REGION Network 5: Estado 3
   RUNG wire#powerrail
      { S7_Templates := "SrcType := DWord" } EQ_Contact(in1 := #Prioritaria, in2 := 16#0000_0000)
      { S7_Templates := "SrcType := DWord" } EQ_Contact(in1 := #Concatenadora, in2 := 16#0000_0004)
      wire#w1
      I_Contact( #"Falla Prioritarias" )
      I_Contact( #"Error Concatenadoras" )
      { S7_GenerateENO := "TRUE" } Move(in := 16#0000_0004, out1 => #Estado)
   END_RUNG
   RUNG wire#powerrail
      { S7_Templates := "SrcType := DWord" } EQ_Contact(in1 := #Prioritaria, in2 := 16#0000_0004)
   END_RUNG wire#w1
   // the same network as SCL:
   IF (((#Prioritaria = 16#0000_0000) AND (#Concatenadora = 16#0000_0004)) OR (#Prioritaria = 16#0000_0004)) AND NOT #"Falla Prioritarias" AND NOT #"Error Concatenadoras" THEN
       #Estado := 16#0000_0004;
   END_IF;
END_REGION

REGION Network 6: Estado 4
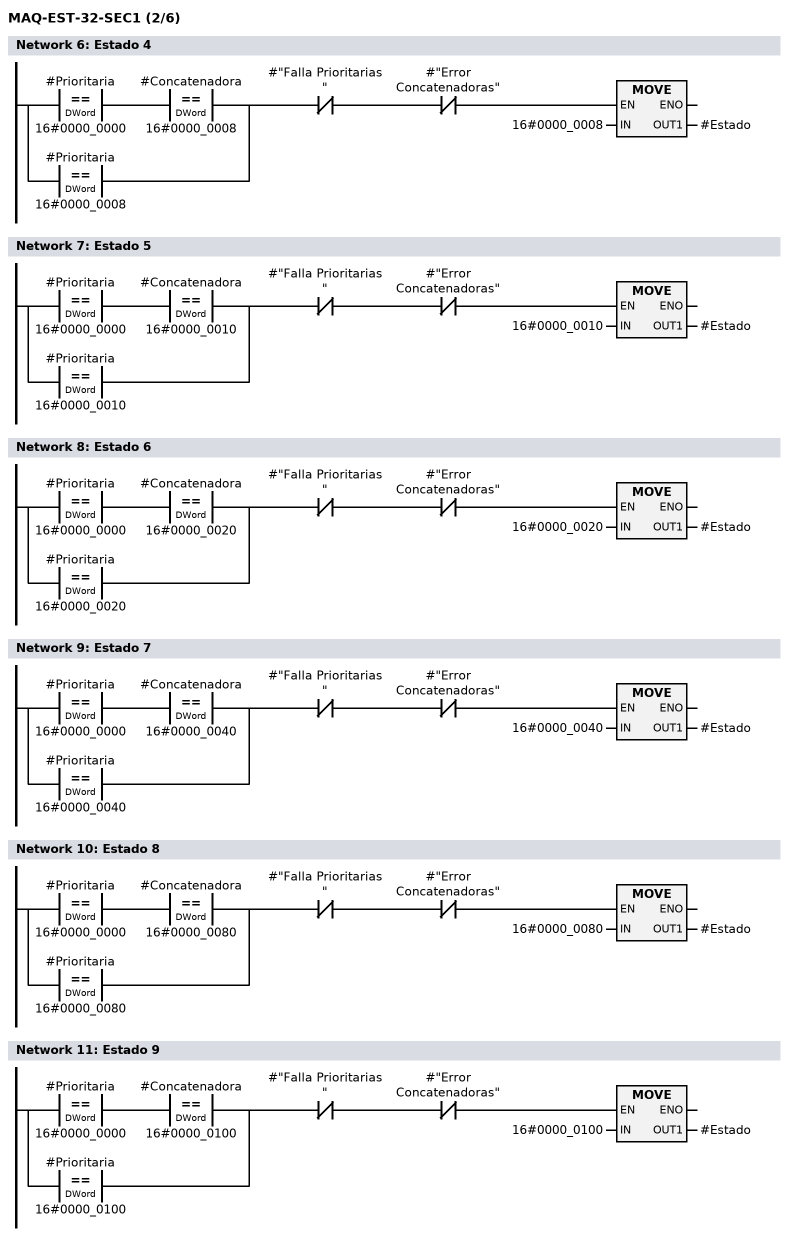
   RUNG wire#powerrail
      { S7_Templates := "SrcType := DWord" } EQ_Contact(in1 := #Prioritaria, in2 := 16#0000_0000)
      { S7_Templates := "SrcType := DWord" } EQ_Contact(in1 := #Concatenadora, in2 := 16#0000_0008)
      wire#w1
      I_Contact( #"Falla Prioritarias" )
      I_Contact( #"Error Concatenadoras" )
      { S7_GenerateENO := "TRUE" } Move(in := 16#0000_0008, out1 => #Estado)
   END_RUNG
   RUNG wire#powerrail
      { S7_Templates := "SrcType := DWord" } EQ_Contact(in1 := #Prioritaria, in2 := 16#0000_0008)
   END_RUNG wire#w1
   // the same network as SCL:
   IF (((#Prioritaria = 16#0000_0000) AND (#Concatenadora = 16#0000_0008)) OR (#Prioritaria = 16#0000_0008)) AND NOT #"Falla Prioritarias" AND NOT #"Error Concatenadoras" THEN
       #Estado := 16#0000_0008;
   END_IF;
END_REGION

REGION Network 7: Estado 5
   RUNG wire#powerrail
      { S7_Templates := "SrcType := DWord" } EQ_Contact(in1 := #Prioritaria, in2 := 16#0000_0000)
      { S7_Templates := "SrcType := DWord" } EQ_Contact(in1 := #Concatenadora, in2 := 16#0000_0010)
      wire#w1
      I_Contact( #"Falla Prioritarias" )
      I_Contact( #"Error Concatenadoras" )
      { S7_GenerateENO := "TRUE" } Move(in := 16#0000_0010, out1 => #Estado)
   END_RUNG
   RUNG wire#powerrail
      { S7_Templates := "SrcType := DWord" } EQ_Contact(in1 := #Prioritaria, in2 := 16#0000_0010)
   END_RUNG wire#w1
   // the same network as SCL:
   IF (((#Prioritaria = 16#0000_0000) AND (#Concatenadora = 16#0000_0010)) OR (#Prioritaria = 16#0000_0010)) AND NOT #"Falla Prioritarias" AND NOT #"Error Concatenadoras" THEN
       #Estado := 16#0000_0010;
   END_IF;
END_REGION

REGION Network 8: Estado 6
   RUNG wire#powerrail
      { S7_Templates := "SrcType := DWord" } EQ_Contact(in1 := #Prioritaria, in2 := 16#0000_0000)
      { S7_Templates := "SrcType := DWord" } EQ_Contact(in1 := #Concatenadora, in2 := 16#0000_0020)
      wire#w1
      I_Contact( #"Falla Prioritarias" )
      I_Contact( #"Error Concatenadoras" )
      { S7_GenerateENO := "TRUE" } Move(in := 16#0000_0020, out1 => #Estado)
   END_RUNG
   RUNG wire#powerrail
      { S7_Templates := "SrcType := DWord" } EQ_Contact(in1 := #Prioritaria, in2 := 16#0000_0020)
   END_RUNG wire#w1
   // the same network as SCL:
   IF (((#Prioritaria = 16#0000_0000) AND (#Concatenadora = 16#0000_0020)) OR (#Prioritaria = 16#0000_0020)) AND NOT #"Falla Prioritarias" AND NOT #"Error Concatenadoras" THEN
       #Estado := 16#0000_0020;
   END_IF;
END_REGION

REGION Network 9: Estado 7
   RUNG wire#powerrail
      { S7_Templates := "SrcType := DWord" } EQ_Contact(in1 := #Prioritaria, in2 := 16#0000_0000)
      { S7_Templates := "SrcType := DWord" } EQ_Contact(in1 := #Concatenadora, in2 := 16#0000_0040)
      wire#w1
      I_Contact( #"Falla Prioritarias" )
      I_Contact( #"Error Concatenadoras" )
      { S7_GenerateENO := "TRUE" } Move(in := 16#0000_0040, out1 => #Estado)
   END_RUNG
   RUNG wire#powerrail
      { S7_Templates := "SrcType := DWord" } EQ_Contact(in1 := #Prioritaria, in2 := 16#0000_0040)
   END_RUNG wire#w1
   // the same network as SCL:
   IF (((#Prioritaria = 16#0000_0000) AND (#Concatenadora = 16#0000_0040)) OR (#Prioritaria = 16#0000_0040)) AND NOT #"Falla Prioritarias" AND NOT #"Error Concatenadoras" THEN
       #Estado := 16#0000_0040;
   END_IF;
END_REGION

REGION Network 10: Estado 8
   RUNG wire#powerrail
      { S7_Templates := "SrcType := DWord" } EQ_Contact(in1 := #Prioritaria, in2 := 16#0000_0000)
      { S7_Templates := "SrcType := DWord" } EQ_Contact(in1 := #Concatenadora, in2 := 16#0000_0080)
      wire#w1
      I_Contact( #"Falla Prioritarias" )
      I_Contact( #"Error Concatenadoras" )
      { S7_GenerateENO := "TRUE" } Move(in := 16#0000_0080, out1 => #Estado)
   END_RUNG
   RUNG wire#powerrail
      { S7_Templates := "SrcType := DWord" } EQ_Contact(in1 := #Prioritaria, in2 := 16#0000_0080)
   END_RUNG wire#w1
   // the same network as SCL:
   IF (((#Prioritaria = 16#0000_0000) AND (#Concatenadora = 16#0000_0080)) OR (#Prioritaria = 16#0000_0080)) AND NOT #"Falla Prioritarias" AND NOT #"Error Concatenadoras" THEN
       #Estado := 16#0000_0080;
   END_IF;
END_REGION

REGION Network 11: Estado 9
   RUNG wire#powerrail
      { S7_Templates := "SrcType := DWord" } EQ_Contact(in1 := #Prioritaria, in2 := 16#0000_0000)
      { S7_Templates := "SrcType := DWord" } EQ_Contact(in1 := #Concatenadora, in2 := 16#0000_0100)
      wire#w1
      I_Contact( #"Falla Prioritarias" )
      I_Contact( #"Error Concatenadoras" )
      { S7_GenerateENO := "TRUE" } Move(in := 16#0000_0100, out1 => #Estado)
   END_RUNG
   RUNG wire#powerrail
      { S7_Templates := "SrcType := DWord" } EQ_Contact(in1 := #Prioritaria, in2 := 16#0000_0100)
   END_RUNG wire#w1
   // the same network as SCL:
   IF (((#Prioritaria = 16#0000_0000) AND (#Concatenadora = 16#0000_0100)) OR (#Prioritaria = 16#0000_0100)) AND NOT #"Falla Prioritarias" AND NOT #"Error Concatenadoras" THEN
       #Estado := 16#0000_0100;
   END_IF;
END_REGION

REGION Network 12: Estado 10
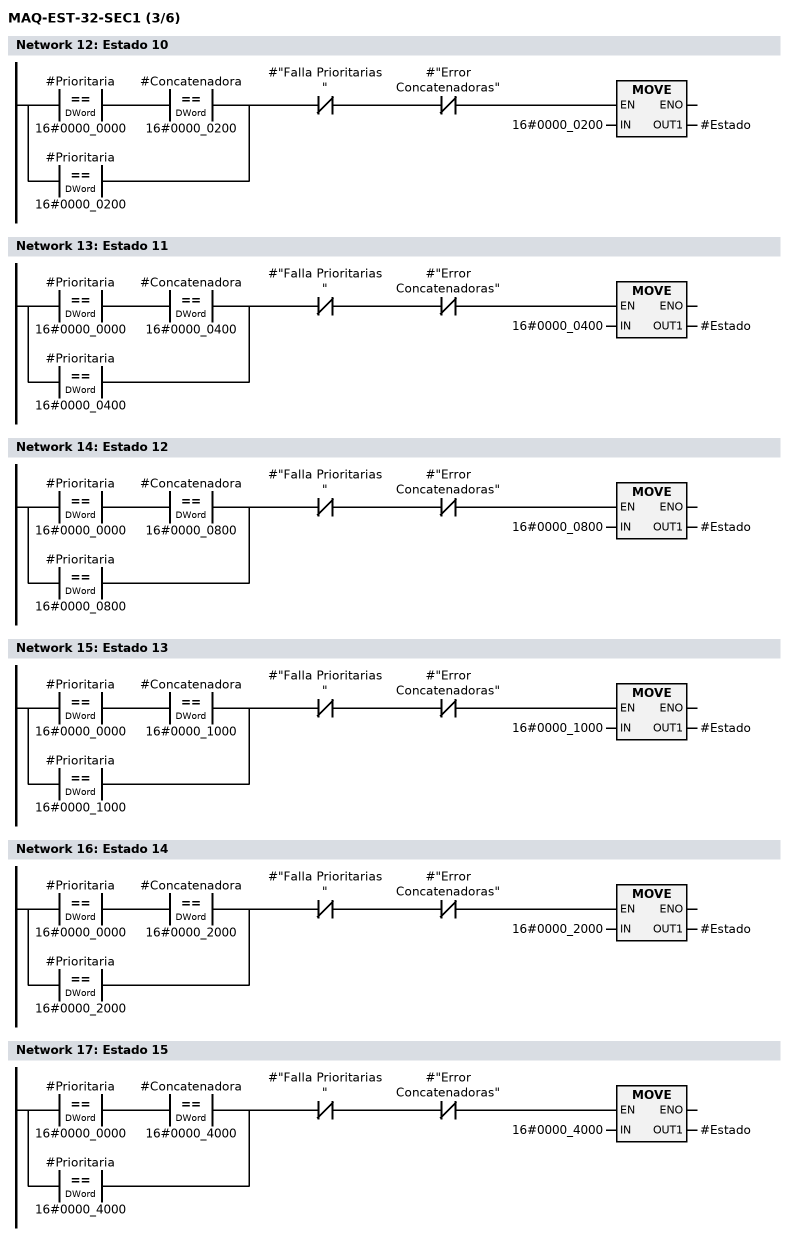
   RUNG wire#powerrail
      { S7_Templates := "SrcType := DWord" } EQ_Contact(in1 := #Prioritaria, in2 := 16#0000_0000)
      { S7_Templates := "SrcType := DWord" } EQ_Contact(in1 := #Concatenadora, in2 := 16#0000_0200)
      wire#w1
      I_Contact( #"Falla Prioritarias" )
      I_Contact( #"Error Concatenadoras" )
      { S7_GenerateENO := "TRUE" } Move(in := 16#0000_0200, out1 => #Estado)
   END_RUNG
   RUNG wire#powerrail
      { S7_Templates := "SrcType := DWord" } EQ_Contact(in1 := #Prioritaria, in2 := 16#0000_0200)
   END_RUNG wire#w1
   // the same network as SCL:
   IF (((#Prioritaria = 16#0000_0000) AND (#Concatenadora = 16#0000_0200)) OR (#Prioritaria = 16#0000_0200)) AND NOT #"Falla Prioritarias" AND NOT #"Error Concatenadoras" THEN
       #Estado := 16#0000_0200;
   END_IF;
END_REGION

REGION Network 13: Estado 11
   RUNG wire#powerrail
      { S7_Templates := "SrcType := DWord" } EQ_Contact(in1 := #Prioritaria, in2 := 16#0000_0000)
      { S7_Templates := "SrcType := DWord" } EQ_Contact(in1 := #Concatenadora, in2 := 16#0000_0400)
      wire#w1
      I_Contact( #"Falla Prioritarias" )
      I_Contact( #"Error Concatenadoras" )
      { S7_GenerateENO := "TRUE" } Move(in := 16#0000_0400, out1 => #Estado)
   END_RUNG
   RUNG wire#powerrail
      { S7_Templates := "SrcType := DWord" } EQ_Contact(in1 := #Prioritaria, in2 := 16#0000_0400)
   END_RUNG wire#w1
   // the same network as SCL:
   IF (((#Prioritaria = 16#0000_0000) AND (#Concatenadora = 16#0000_0400)) OR (#Prioritaria = 16#0000_0400)) AND NOT #"Falla Prioritarias" AND NOT #"Error Concatenadoras" THEN
       #Estado := 16#0000_0400;
   END_IF;
END_REGION

REGION Network 14: Estado 12
   RUNG wire#powerrail
      { S7_Templates := "SrcType := DWord" } EQ_Contact(in1 := #Prioritaria, in2 := 16#0000_0000)
      { S7_Templates := "SrcType := DWord" } EQ_Contact(in1 := #Concatenadora, in2 := 16#0000_0800)
      wire#w1
      I_Contact( #"Falla Prioritarias" )
      I_Contact( #"Error Concatenadoras" )
      { S7_GenerateENO := "TRUE" } Move(in := 16#0000_0800, out1 => #Estado)
   END_RUNG
   RUNG wire#powerrail
      { S7_Templates := "SrcType := DWord" } EQ_Contact(in1 := #Prioritaria, in2 := 16#0000_0800)
   END_RUNG wire#w1
   // the same network as SCL:
   IF (((#Prioritaria = 16#0000_0000) AND (#Concatenadora = 16#0000_0800)) OR (#Prioritaria = 16#0000_0800)) AND NOT #"Falla Prioritarias" AND NOT #"Error Concatenadoras" THEN
       #Estado := 16#0000_0800;
   END_IF;
END_REGION

REGION Network 15: Estado 13
   RUNG wire#powerrail
      { S7_Templates := "SrcType := DWord" } EQ_Contact(in1 := #Prioritaria, in2 := 16#0000_0000)
      { S7_Templates := "SrcType := DWord" } EQ_Contact(in1 := #Concatenadora, in2 := 16#0000_1000)
      wire#w1
      I_Contact( #"Falla Prioritarias" )
      I_Contact( #"Error Concatenadoras" )
      { S7_GenerateENO := "TRUE" } Move(in := 16#0000_1000, out1 => #Estado)
   END_RUNG
   RUNG wire#powerrail
      { S7_Templates := "SrcType := DWord" } EQ_Contact(in1 := #Prioritaria, in2 := 16#0000_1000)
   END_RUNG wire#w1
   // the same network as SCL:
   IF (((#Prioritaria = 16#0000_0000) AND (#Concatenadora = 16#0000_1000)) OR (#Prioritaria = 16#0000_1000)) AND NOT #"Falla Prioritarias" AND NOT #"Error Concatenadoras" THEN
       #Estado := 16#0000_1000;
   END_IF;
END_REGION

REGION Network 16: Estado 14
   RUNG wire#powerrail
      { S7_Templates := "SrcType := DWord" } EQ_Contact(in1 := #Prioritaria, in2 := 16#0000_0000)
      { S7_Templates := "SrcType := DWord" } EQ_Contact(in1 := #Concatenadora, in2 := 16#0000_2000)
      wire#w1
      I_Contact( #"Falla Prioritarias" )
      I_Contact( #"Error Concatenadoras" )
      { S7_GenerateENO := "TRUE" } Move(in := 16#0000_2000, out1 => #Estado)
   END_RUNG
   RUNG wire#powerrail
      { S7_Templates := "SrcType := DWord" } EQ_Contact(in1 := #Prioritaria, in2 := 16#0000_2000)
   END_RUNG wire#w1
   // the same network as SCL:
   IF (((#Prioritaria = 16#0000_0000) AND (#Concatenadora = 16#0000_2000)) OR (#Prioritaria = 16#0000_2000)) AND NOT #"Falla Prioritarias" AND NOT #"Error Concatenadoras" THEN
       #Estado := 16#0000_2000;
   END_IF;
END_REGION

REGION Network 17: Estado 15
   RUNG wire#powerrail
      { S7_Templates := "SrcType := DWord" } EQ_Contact(in1 := #Prioritaria, in2 := 16#0000_0000)
      { S7_Templates := "SrcType := DWord" } EQ_Contact(in1 := #Concatenadora, in2 := 16#0000_4000)
      wire#w1
      I_Contact( #"Falla Prioritarias" )
      I_Contact( #"Error Concatenadoras" )
      { S7_GenerateENO := "TRUE" } Move(in := 16#0000_4000, out1 => #Estado)
   END_RUNG
   RUNG wire#powerrail
      { S7_Templates := "SrcType := DWord" } EQ_Contact(in1 := #Prioritaria, in2 := 16#0000_4000)
   END_RUNG wire#w1
   // the same network as SCL:
   IF (((#Prioritaria = 16#0000_0000) AND (#Concatenadora = 16#0000_4000)) OR (#Prioritaria = 16#0000_4000)) AND NOT #"Falla Prioritarias" AND NOT #"Error Concatenadoras" THEN
       #Estado := 16#0000_4000;
   END_IF;
END_REGION

REGION Network 18: Estado 16
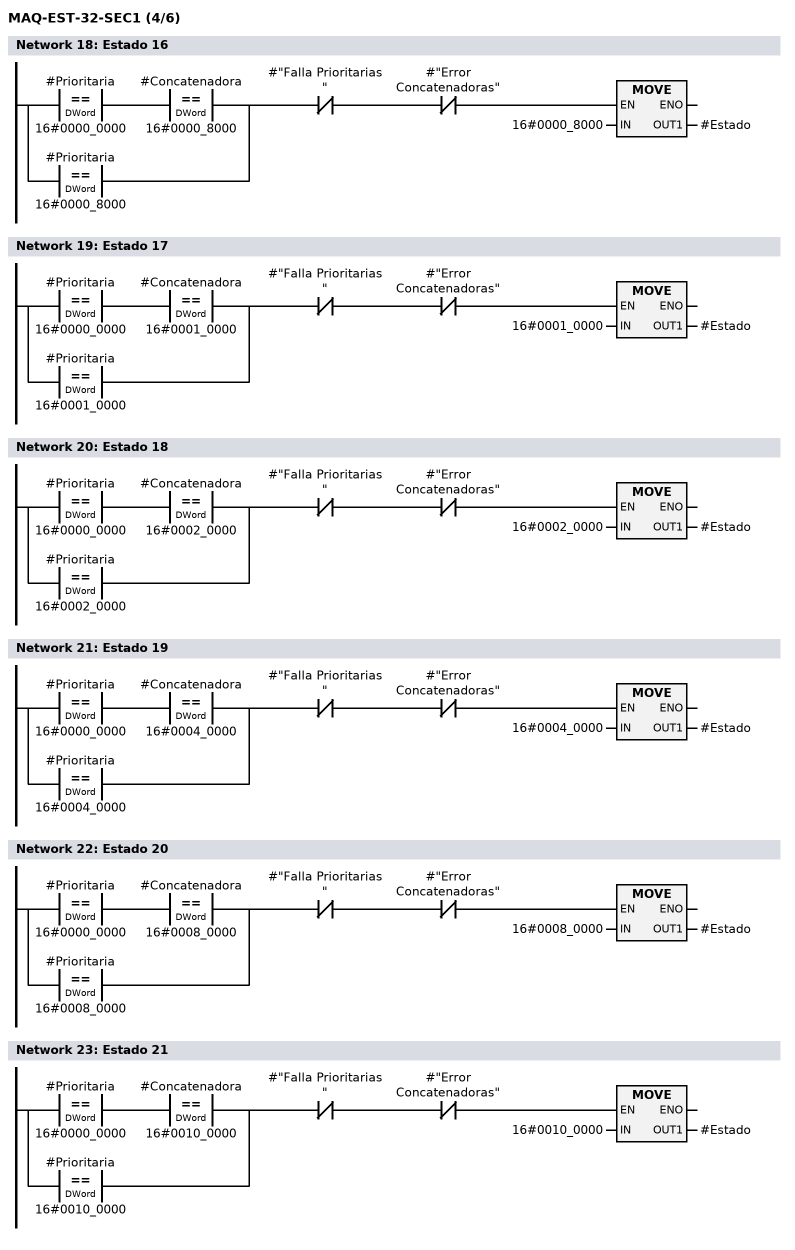
   RUNG wire#powerrail
      { S7_Templates := "SrcType := DWord" } EQ_Contact(in1 := #Prioritaria, in2 := 16#0000_0000)
      { S7_Templates := "SrcType := DWord" } EQ_Contact(in1 := #Concatenadora, in2 := 16#0000_8000)
      wire#w1
      I_Contact( #"Falla Prioritarias" )
      I_Contact( #"Error Concatenadoras" )
      { S7_GenerateENO := "TRUE" } Move(in := 16#0000_8000, out1 => #Estado)
   END_RUNG
   RUNG wire#powerrail
      { S7_Templates := "SrcType := DWord" } EQ_Contact(in1 := #Prioritaria, in2 := 16#0000_8000)
   END_RUNG wire#w1
   // the same network as SCL:
   IF (((#Prioritaria = 16#0000_0000) AND (#Concatenadora = 16#0000_8000)) OR (#Prioritaria = 16#0000_8000)) AND NOT #"Falla Prioritarias" AND NOT #"Error Concatenadoras" THEN
       #Estado := 16#0000_8000;
   END_IF;
END_REGION

REGION Network 19: Estado 17
   RUNG wire#powerrail
      { S7_Templates := "SrcType := DWord" } EQ_Contact(in1 := #Prioritaria, in2 := 16#0000_0000)
      { S7_Templates := "SrcType := DWord" } EQ_Contact(in1 := #Concatenadora, in2 := 16#0001_0000)
      wire#w1
      I_Contact( #"Falla Prioritarias" )
      I_Contact( #"Error Concatenadoras" )
      { S7_GenerateENO := "TRUE" } Move(in := 16#0001_0000, out1 => #Estado)
   END_RUNG
   RUNG wire#powerrail
      { S7_Templates := "SrcType := DWord" } EQ_Contact(in1 := #Prioritaria, in2 := 16#0001_0000)
   END_RUNG wire#w1
   // the same network as SCL:
   IF (((#Prioritaria = 16#0000_0000) AND (#Concatenadora = 16#0001_0000)) OR (#Prioritaria = 16#0001_0000)) AND NOT #"Falla Prioritarias" AND NOT #"Error Concatenadoras" THEN
       #Estado := 16#0001_0000;
   END_IF;
END_REGION

REGION Network 20: Estado 18
   RUNG wire#powerrail
      { S7_Templates := "SrcType := DWord" } EQ_Contact(in1 := #Prioritaria, in2 := 16#0000_0000)
      { S7_Templates := "SrcType := DWord" } EQ_Contact(in1 := #Concatenadora, in2 := 16#0002_0000)
      wire#w1
      I_Contact( #"Falla Prioritarias" )
      I_Contact( #"Error Concatenadoras" )
      { S7_GenerateENO := "TRUE" } Move(in := 16#0002_0000, out1 => #Estado)
   END_RUNG
   RUNG wire#powerrail
      { S7_Templates := "SrcType := DWord" } EQ_Contact(in1 := #Prioritaria, in2 := 16#0002_0000)
   END_RUNG wire#w1
   // the same network as SCL:
   IF (((#Prioritaria = 16#0000_0000) AND (#Concatenadora = 16#0002_0000)) OR (#Prioritaria = 16#0002_0000)) AND NOT #"Falla Prioritarias" AND NOT #"Error Concatenadoras" THEN
       #Estado := 16#0002_0000;
   END_IF;
END_REGION

REGION Network 21: Estado 19
   RUNG wire#powerrail
      { S7_Templates := "SrcType := DWord" } EQ_Contact(in1 := #Prioritaria, in2 := 16#0000_0000)
      { S7_Templates := "SrcType := DWord" } EQ_Contact(in1 := #Concatenadora, in2 := 16#0004_0000)
      wire#w1
      I_Contact( #"Falla Prioritarias" )
      I_Contact( #"Error Concatenadoras" )
      { S7_GenerateENO := "TRUE" } Move(in := 16#0004_0000, out1 => #Estado)
   END_RUNG
   RUNG wire#powerrail
      { S7_Templates := "SrcType := DWord" } EQ_Contact(in1 := #Prioritaria, in2 := 16#0004_0000)
   END_RUNG wire#w1
   // the same network as SCL:
   IF (((#Prioritaria = 16#0000_0000) AND (#Concatenadora = 16#0004_0000)) OR (#Prioritaria = 16#0004_0000)) AND NOT #"Falla Prioritarias" AND NOT #"Error Concatenadoras" THEN
       #Estado := 16#0004_0000;
   END_IF;
END_REGION

REGION Network 22: Estado 20
   RUNG wire#powerrail
      { S7_Templates := "SrcType := DWord" } EQ_Contact(in1 := #Prioritaria, in2 := 16#0000_0000)
      { S7_Templates := "SrcType := DWord" } EQ_Contact(in1 := #Concatenadora, in2 := 16#0008_0000)
      wire#w1
      I_Contact( #"Falla Prioritarias" )
      I_Contact( #"Error Concatenadoras" )
      { S7_GenerateENO := "TRUE" } Move(in := 16#0008_0000, out1 => #Estado)
   END_RUNG
   RUNG wire#powerrail
      { S7_Templates := "SrcType := DWord" } EQ_Contact(in1 := #Prioritaria, in2 := 16#0008_0000)
   END_RUNG wire#w1
   // the same network as SCL:
   IF (((#Prioritaria = 16#0000_0000) AND (#Concatenadora = 16#0008_0000)) OR (#Prioritaria = 16#0008_0000)) AND NOT #"Falla Prioritarias" AND NOT #"Error Concatenadoras" THEN
       #Estado := 16#0008_0000;
   END_IF;
END_REGION

REGION Network 23: Estado 21
   RUNG wire#powerrail
      { S7_Templates := "SrcType := DWord" } EQ_Contact(in1 := #Prioritaria, in2 := 16#0000_0000)
      { S7_Templates := "SrcType := DWord" } EQ_Contact(in1 := #Concatenadora, in2 := 16#0010_0000)
      wire#w1
      I_Contact( #"Falla Prioritarias" )
      I_Contact( #"Error Concatenadoras" )
      { S7_GenerateENO := "TRUE" } Move(in := 16#0010_0000, out1 => #Estado)
   END_RUNG
   RUNG wire#powerrail
      { S7_Templates := "SrcType := DWord" } EQ_Contact(in1 := #Prioritaria, in2 := 16#0010_0000)
   END_RUNG wire#w1
   // the same network as SCL:
   IF (((#Prioritaria = 16#0000_0000) AND (#Concatenadora = 16#0010_0000)) OR (#Prioritaria = 16#0010_0000)) AND NOT #"Falla Prioritarias" AND NOT #"Error Concatenadoras" THEN
       #Estado := 16#0010_0000;
   END_IF;
END_REGION

REGION Network 24: Estado 22
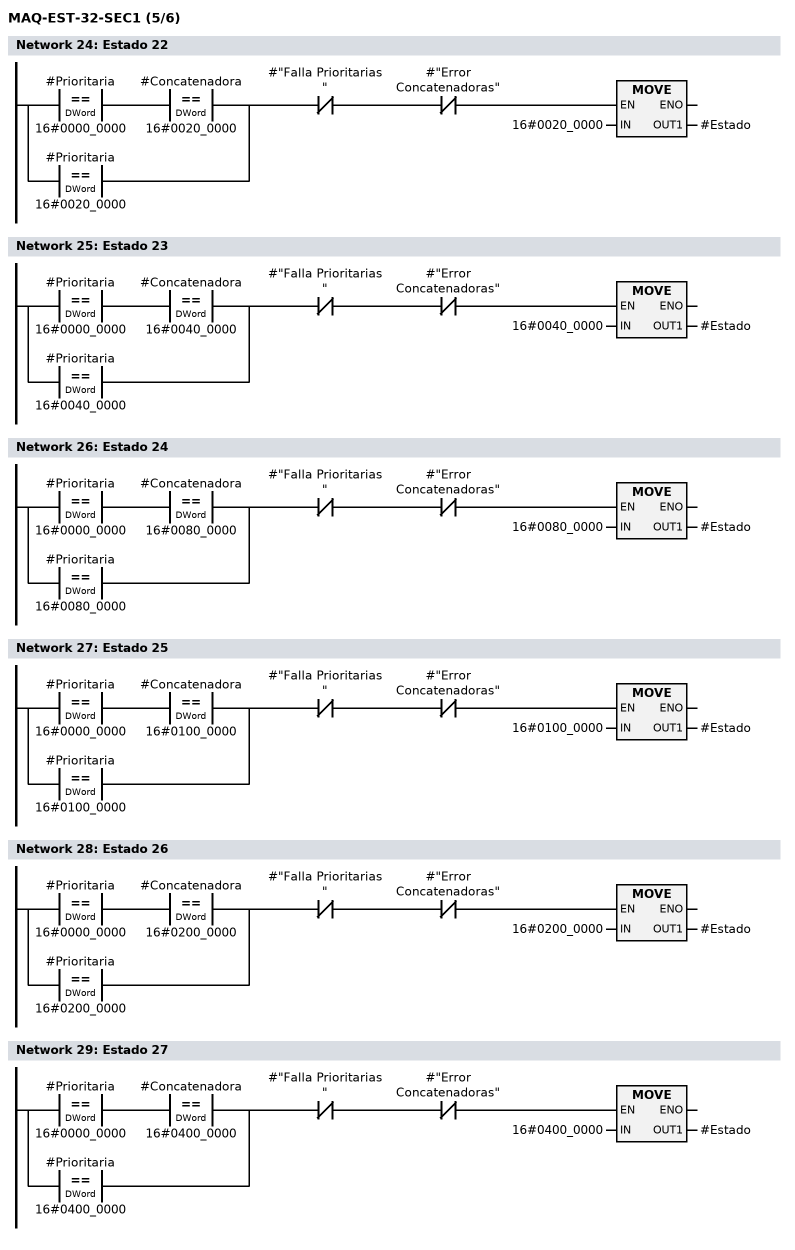
   RUNG wire#powerrail
      { S7_Templates := "SrcType := DWord" } EQ_Contact(in1 := #Prioritaria, in2 := 16#0000_0000)
      { S7_Templates := "SrcType := DWord" } EQ_Contact(in1 := #Concatenadora, in2 := 16#0020_0000)
      wire#w1
      I_Contact( #"Falla Prioritarias" )
      I_Contact( #"Error Concatenadoras" )
      { S7_GenerateENO := "TRUE" } Move(in := 16#0020_0000, out1 => #Estado)
   END_RUNG
   RUNG wire#powerrail
      { S7_Templates := "SrcType := DWord" } EQ_Contact(in1 := #Prioritaria, in2 := 16#0020_0000)
   END_RUNG wire#w1
   // the same network as SCL:
   IF (((#Prioritaria = 16#0000_0000) AND (#Concatenadora = 16#0020_0000)) OR (#Prioritaria = 16#0020_0000)) AND NOT #"Falla Prioritarias" AND NOT #"Error Concatenadoras" THEN
       #Estado := 16#0020_0000;
   END_IF;
END_REGION

REGION Network 25: Estado 23
   RUNG wire#powerrail
      { S7_Templates := "SrcType := DWord" } EQ_Contact(in1 := #Prioritaria, in2 := 16#0000_0000)
      { S7_Templates := "SrcType := DWord" } EQ_Contact(in1 := #Concatenadora, in2 := 16#0040_0000)
      wire#w1
      I_Contact( #"Falla Prioritarias" )
      I_Contact( #"Error Concatenadoras" )
      { S7_GenerateENO := "TRUE" } Move(in := 16#0040_0000, out1 => #Estado)
   END_RUNG
   RUNG wire#powerrail
      { S7_Templates := "SrcType := DWord" } EQ_Contact(in1 := #Prioritaria, in2 := 16#0040_0000)
   END_RUNG wire#w1
   // the same network as SCL:
   IF (((#Prioritaria = 16#0000_0000) AND (#Concatenadora = 16#0040_0000)) OR (#Prioritaria = 16#0040_0000)) AND NOT #"Falla Prioritarias" AND NOT #"Error Concatenadoras" THEN
       #Estado := 16#0040_0000;
   END_IF;
END_REGION

REGION Network 26: Estado 24
   RUNG wire#powerrail
      { S7_Templates := "SrcType := DWord" } EQ_Contact(in1 := #Prioritaria, in2 := 16#0000_0000)
      { S7_Templates := "SrcType := DWord" } EQ_Contact(in1 := #Concatenadora, in2 := 16#0080_0000)
      wire#w1
      I_Contact( #"Falla Prioritarias" )
      I_Contact( #"Error Concatenadoras" )
      { S7_GenerateENO := "TRUE" } Move(in := 16#0080_0000, out1 => #Estado)
   END_RUNG
   RUNG wire#powerrail
      { S7_Templates := "SrcType := DWord" } EQ_Contact(in1 := #Prioritaria, in2 := 16#0080_0000)
   END_RUNG wire#w1
   // the same network as SCL:
   IF (((#Prioritaria = 16#0000_0000) AND (#Concatenadora = 16#0080_0000)) OR (#Prioritaria = 16#0080_0000)) AND NOT #"Falla Prioritarias" AND NOT #"Error Concatenadoras" THEN
       #Estado := 16#0080_0000;
   END_IF;
END_REGION

REGION Network 27: Estado 25
   RUNG wire#powerrail
      { S7_Templates := "SrcType := DWord" } EQ_Contact(in1 := #Prioritaria, in2 := 16#0000_0000)
      { S7_Templates := "SrcType := DWord" } EQ_Contact(in1 := #Concatenadora, in2 := 16#0100_0000)
      wire#w1
      I_Contact( #"Falla Prioritarias" )
      I_Contact( #"Error Concatenadoras" )
      { S7_GenerateENO := "TRUE" } Move(in := 16#0100_0000, out1 => #Estado)
   END_RUNG
   RUNG wire#powerrail
      { S7_Templates := "SrcType := DWord" } EQ_Contact(in1 := #Prioritaria, in2 := 16#0100_0000)
   END_RUNG wire#w1
   // the same network as SCL:
   IF (((#Prioritaria = 16#0000_0000) AND (#Concatenadora = 16#0100_0000)) OR (#Prioritaria = 16#0100_0000)) AND NOT #"Falla Prioritarias" AND NOT #"Error Concatenadoras" THEN
       #Estado := 16#0100_0000;
   END_IF;
END_REGION

REGION Network 28: Estado 26
   RUNG wire#powerrail
      { S7_Templates := "SrcType := DWord" } EQ_Contact(in1 := #Prioritaria, in2 := 16#0000_0000)
      { S7_Templates := "SrcType := DWord" } EQ_Contact(in1 := #Concatenadora, in2 := 16#0200_0000)
      wire#w1
      I_Contact( #"Falla Prioritarias" )
      I_Contact( #"Error Concatenadoras" )
      { S7_GenerateENO := "TRUE" } Move(in := 16#0200_0000, out1 => #Estado)
   END_RUNG
   RUNG wire#powerrail
      { S7_Templates := "SrcType := DWord" } EQ_Contact(in1 := #Prioritaria, in2 := 16#0200_0000)
   END_RUNG wire#w1
   // the same network as SCL:
   IF (((#Prioritaria = 16#0000_0000) AND (#Concatenadora = 16#0200_0000)) OR (#Prioritaria = 16#0200_0000)) AND NOT #"Falla Prioritarias" AND NOT #"Error Concatenadoras" THEN
       #Estado := 16#0200_0000;
   END_IF;
END_REGION

REGION Network 29: Estado 27
   RUNG wire#powerrail
      { S7_Templates := "SrcType := DWord" } EQ_Contact(in1 := #Prioritaria, in2 := 16#0000_0000)
      { S7_Templates := "SrcType := DWord" } EQ_Contact(in1 := #Concatenadora, in2 := 16#0400_0000)
      wire#w1
      I_Contact( #"Falla Prioritarias" )
      I_Contact( #"Error Concatenadoras" )
      { S7_GenerateENO := "TRUE" } Move(in := 16#0400_0000, out1 => #Estado)
   END_RUNG
   RUNG wire#powerrail
      { S7_Templates := "SrcType := DWord" } EQ_Contact(in1 := #Prioritaria, in2 := 16#0400_0000)
   END_RUNG wire#w1
   // the same network as SCL:
   IF (((#Prioritaria = 16#0000_0000) AND (#Concatenadora = 16#0400_0000)) OR (#Prioritaria = 16#0400_0000)) AND NOT #"Falla Prioritarias" AND NOT #"Error Concatenadoras" THEN
       #Estado := 16#0400_0000;
   END_IF;
END_REGION

REGION Network 30: Estado 28
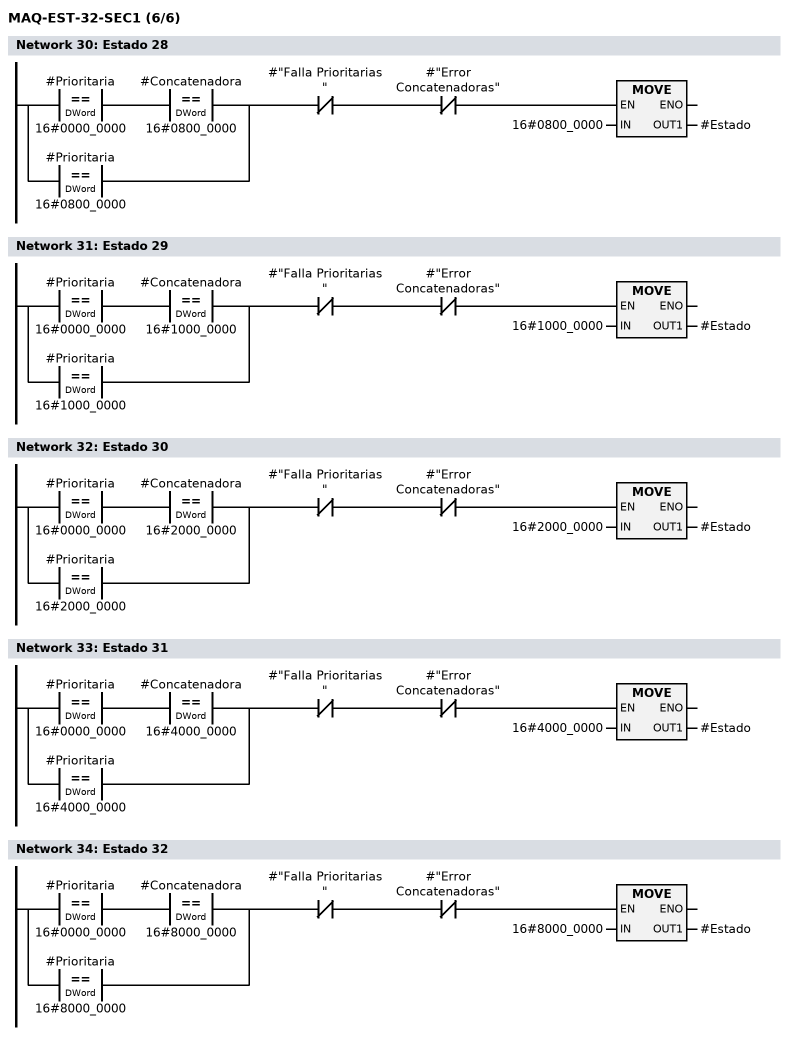
   RUNG wire#powerrail
      { S7_Templates := "SrcType := DWord" } EQ_Contact(in1 := #Prioritaria, in2 := 16#0000_0000)
      { S7_Templates := "SrcType := DWord" } EQ_Contact(in1 := #Concatenadora, in2 := 16#0800_0000)
      wire#w1
      I_Contact( #"Falla Prioritarias" )
      I_Contact( #"Error Concatenadoras" )
      { S7_GenerateENO := "TRUE" } Move(in := 16#0800_0000, out1 => #Estado)
   END_RUNG
   RUNG wire#powerrail
      { S7_Templates := "SrcType := DWord" } EQ_Contact(in1 := #Prioritaria, in2 := 16#0800_0000)
   END_RUNG wire#w1
   // the same network as SCL:
   IF (((#Prioritaria = 16#0000_0000) AND (#Concatenadora = 16#0800_0000)) OR (#Prioritaria = 16#0800_0000)) AND NOT #"Falla Prioritarias" AND NOT #"Error Concatenadoras" THEN
       #Estado := 16#0800_0000;
   END_IF;
END_REGION

REGION Network 31: Estado 29
   RUNG wire#powerrail
      { S7_Templates := "SrcType := DWord" } EQ_Contact(in1 := #Prioritaria, in2 := 16#0000_0000)
      { S7_Templates := "SrcType := DWord" } EQ_Contact(in1 := #Concatenadora, in2 := 16#1000_0000)
      wire#w1
      I_Contact( #"Falla Prioritarias" )
      I_Contact( #"Error Concatenadoras" )
      { S7_GenerateENO := "TRUE" } Move(in := 16#1000_0000, out1 => #Estado)
   END_RUNG
   RUNG wire#powerrail
      { S7_Templates := "SrcType := DWord" } EQ_Contact(in1 := #Prioritaria, in2 := 16#1000_0000)
   END_RUNG wire#w1
   // the same network as SCL:
   IF (((#Prioritaria = 16#0000_0000) AND (#Concatenadora = 16#1000_0000)) OR (#Prioritaria = 16#1000_0000)) AND NOT #"Falla Prioritarias" AND NOT #"Error Concatenadoras" THEN
       #Estado := 16#1000_0000;
   END_IF;
END_REGION

REGION Network 32: Estado 30
   RUNG wire#powerrail
      { S7_Templates := "SrcType := DWord" } EQ_Contact(in1 := #Prioritaria, in2 := 16#0000_0000)
      { S7_Templates := "SrcType := DWord" } EQ_Contact(in1 := #Concatenadora, in2 := 16#2000_0000)
      wire#w1
      I_Contact( #"Falla Prioritarias" )
      I_Contact( #"Error Concatenadoras" )
      { S7_GenerateENO := "TRUE" } Move(in := 16#2000_0000, out1 => #Estado)
   END_RUNG
   RUNG wire#powerrail
      { S7_Templates := "SrcType := DWord" } EQ_Contact(in1 := #Prioritaria, in2 := 16#2000_0000)
   END_RUNG wire#w1
   // the same network as SCL:
   IF (((#Prioritaria = 16#0000_0000) AND (#Concatenadora = 16#2000_0000)) OR (#Prioritaria = 16#2000_0000)) AND NOT #"Falla Prioritarias" AND NOT #"Error Concatenadoras" THEN
       #Estado := 16#2000_0000;
   END_IF;
END_REGION

REGION Network 33: Estado 31
   RUNG wire#powerrail
      { S7_Templates := "SrcType := DWord" } EQ_Contact(in1 := #Prioritaria, in2 := 16#0000_0000)
      { S7_Templates := "SrcType := DWord" } EQ_Contact(in1 := #Concatenadora, in2 := 16#4000_0000)
      wire#w1
      I_Contact( #"Falla Prioritarias" )
      I_Contact( #"Error Concatenadoras" )
      { S7_GenerateENO := "TRUE" } Move(in := 16#4000_0000, out1 => #Estado)
   END_RUNG
   RUNG wire#powerrail
      { S7_Templates := "SrcType := DWord" } EQ_Contact(in1 := #Prioritaria, in2 := 16#4000_0000)
   END_RUNG wire#w1
   // the same network as SCL:
   IF (((#Prioritaria = 16#0000_0000) AND (#Concatenadora = 16#4000_0000)) OR (#Prioritaria = 16#4000_0000)) AND NOT #"Falla Prioritarias" AND NOT #"Error Concatenadoras" THEN
       #Estado := 16#4000_0000;
   END_IF;
END_REGION

REGION Network 34: Estado 32
   RUNG wire#powerrail
      { S7_Templates := "SrcType := DWord" } EQ_Contact(in1 := #Prioritaria, in2 := 16#0000_0000)
      { S7_Templates := "SrcType := DWord" } EQ_Contact(in1 := #Concatenadora, in2 := 16#8000_0000)
      wire#w1
      I_Contact( #"Falla Prioritarias" )
      I_Contact( #"Error Concatenadoras" )
      { S7_GenerateENO := "TRUE" } Move(in := 16#8000_0000, out1 => #Estado)
   END_RUNG
   RUNG wire#powerrail
      { S7_Templates := "SrcType := DWord" } EQ_Contact(in1 := #Prioritaria, in2 := 16#8000_0000)
   END_RUNG wire#w1
   // the same network as SCL:
   IF (((#Prioritaria = 16#0000_0000) AND (#Concatenadora = 16#8000_0000)) OR (#Prioritaria = 16#8000_0000)) AND NOT #"Falla Prioritarias" AND NOT #"Error Concatenadoras" THEN
       #Estado := 16#8000_0000;
   END_IF;
END_REGION
END_FUNCTION

FUNCTION "Brazo de succión" : Void   // FC19, LAD
TITLE = BRAZO DE SUCCIÓN Y BOMBA DE VACÍO.
{ S7_Optimized_Access := 'TRUE' }
VERSION : 0.1
// Es un bloque combinacional que activa el brazo de succión y la bomba, y marca los tiempos del proceso. Hay una marca "ya buscó caja" que indica que el brazo fue arriba a buscar una caja, cuando el brazo baje, y si "busco una caja", activo un temporizador que en el caso que de cumplirse su cuenta, significará que la caja no se desplazó lo suficiente como para permitir que el brazo de succión suba de vuelta. Desde el punto de vista mecánico, el brazo va a estar abajo lo suficiente como para darle tiempo a la cinta a que avance. Es sólo un resguardo. En teoría nunca debería activarse, a menos que haya un problema con la cinta.
   VAR_TEMP   // added for the SCL form of the ladder/FBD networks
      _w1 : Bool;
   END_VAR
BEGIN

REGION Network 1: Activa la bomba
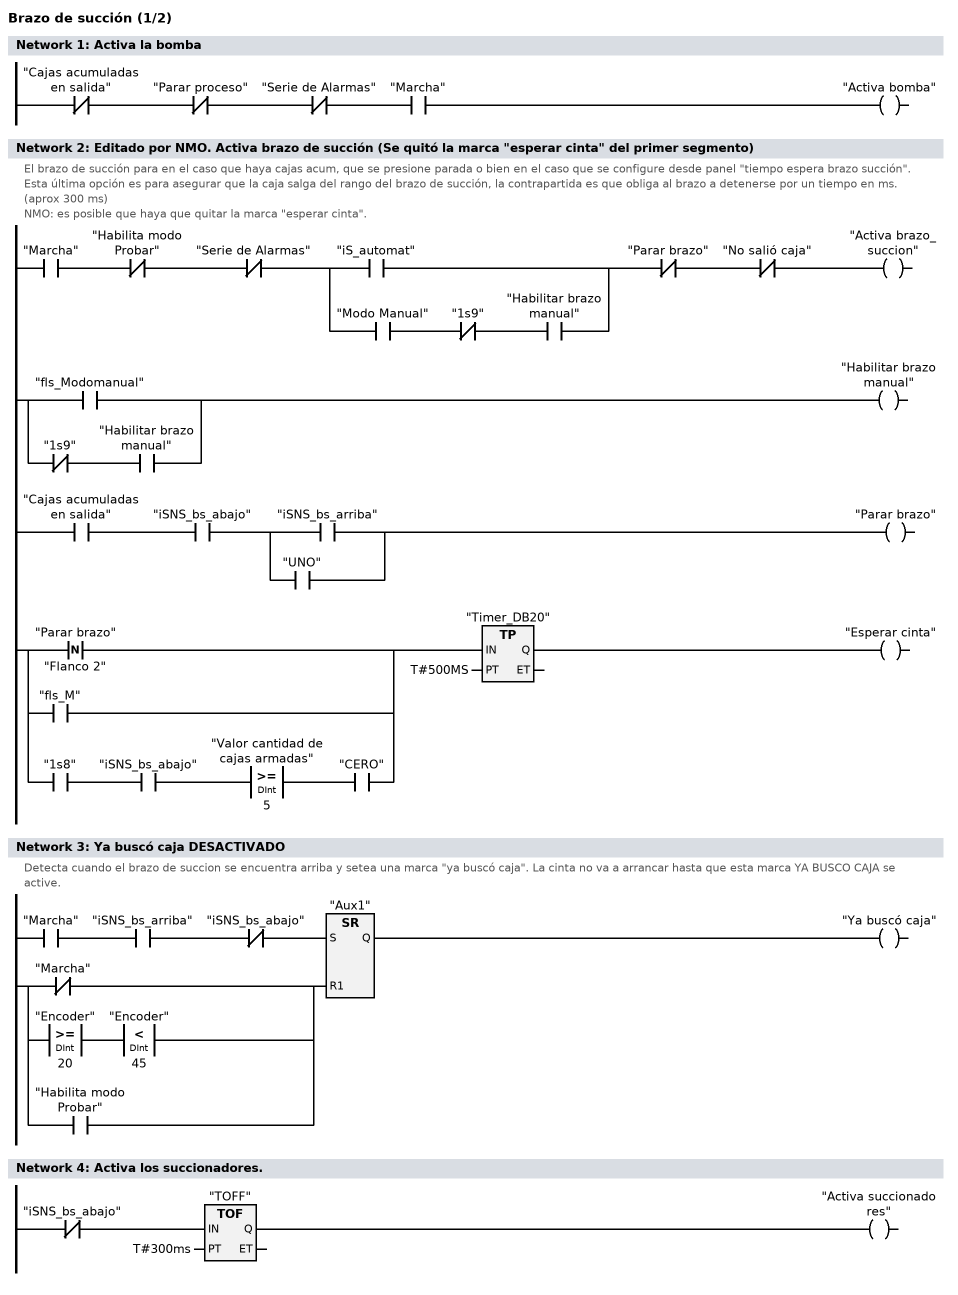
   RUNG wire#powerrail
      I_Contact( "Cajas acumuladas en salida" )
      I_Contact( "Parar proceso" )
      I_Contact( "Serie de Alarmas" )
      Contact( "Marcha" )
      Coil( "Activa bomba" )
   END_RUNG
   // the same network as SCL:
   "Activa bomba" := NOT "Cajas acumuladas en salida" AND NOT "Parar proceso" AND NOT "Serie de Alarmas" AND "Marcha";
END_REGION

REGION Network 2: Editado por NMO. Activa brazo de succión (Se quitó la marca "esperar cinta" del primer segmento)
   // El brazo de succión para en el caso que haya cajas acum, que se presione parada o bien en el caso que se configure desde panel "tiempo espera brazo succión". Esta última opción es para asegurar que la caja salga del rango del brazo de succión, la contrapartida es que obliga al brazo a detenerse por un tiempo en ms. (aprox 300 ms)
   // NMO: es posible que haya que quitar la marca "esperar cinta".
   "Activa brazo_succion" := "Marcha" AND NOT "Habilita modo Probar" AND NOT "Serie de Alarmas" AND ("iS_automat" OR ("Modo Manual" AND NOT "1s9" AND "Habilitar brazo manual")) AND NOT "Parar brazo" AND NOT "No salió caja";
   "Habilitar brazo manual" := "fls_Modomanual" OR (NOT "1s9" AND "Habilitar brazo manual");
   "Parar brazo" := "Cajas acumuladas en salida" AND "iSNS_bs_abajo" AND ("iSNS_bs_arriba" OR "UNO");
   #_w1 := NOT "Parar brazo" AND "Flanco 2";   // falling edge of "Parar brazo"
   "Flanco 2" := "Parar brazo";
   "Timer_DB20".TP(IN := #_w1 OR "fls_M" OR ("1s8" AND "iSNS_bs_abajo" AND ("Valor cantidad de cajas armadas" >= 5) AND "CERO"),
                   PT := T#500MS);
   "Esperar cinta" := "Timer_DB20".Q;
END_REGION
